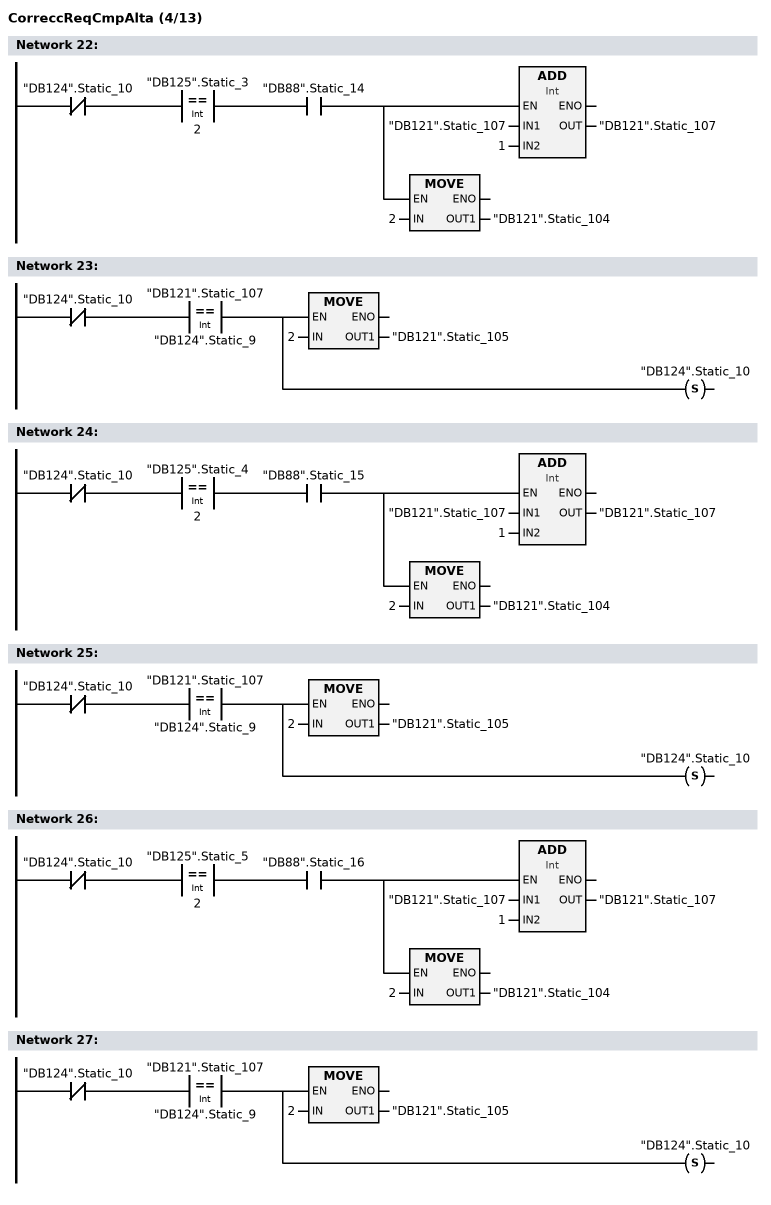
   IF NOT "DB124".Static_10 AND ("DB125".Static_3 = 2) AND "DB88".Static_14 THEN
       "DB121".Static_107 := "DB121".Static_107 + 1;
       "DB121".Static_104 := 2;
   END_IF;
END_REGION

REGION Network 23
   IF NOT "DB124".Static_10 AND ("DB121".Static_107 = "DB124".Static_9) THEN
       "DB121".Static_105 := 2;
       "DB124".Static_10 := TRUE;
   END_IF;
END_REGION

REGION Network 24
   IF NOT "DB124".Static_10 AND ("DB125".Static_4 = 2) AND "DB88".Static_15 THEN
       "DB121".Static_107 := "DB121".Static_107 + 1;
       "DB121".Static_104 := 2;
   END_IF;
END_REGION

REGION Network 25
   IF NOT "DB124".Static_10 AND ("DB121".Static_107 = "DB124".Static_9) THEN
       "DB121".Static_105 := 2;
       "DB124".Static_10 := TRUE;
   END_IF;
END_REGION

REGION Network 26
   IF NOT "DB124".Static_10 AND ("DB125".Static_5 = 2) AND "DB88".Static_16 THEN
       "DB121".Static_107 := "DB121".Static_107 + 1;
       "DB121".Static_104 := 2;
   END_IF;
END_REGION

REGION Network 27
   IF NOT "DB124".Static_10 AND ("DB121".Static_107 = "DB124".Static_9) THEN
       "DB121".Static_105 := 2;
       "DB124".Static_10 := TRUE;
   END_IF;
END_REGION

REGION Network 28
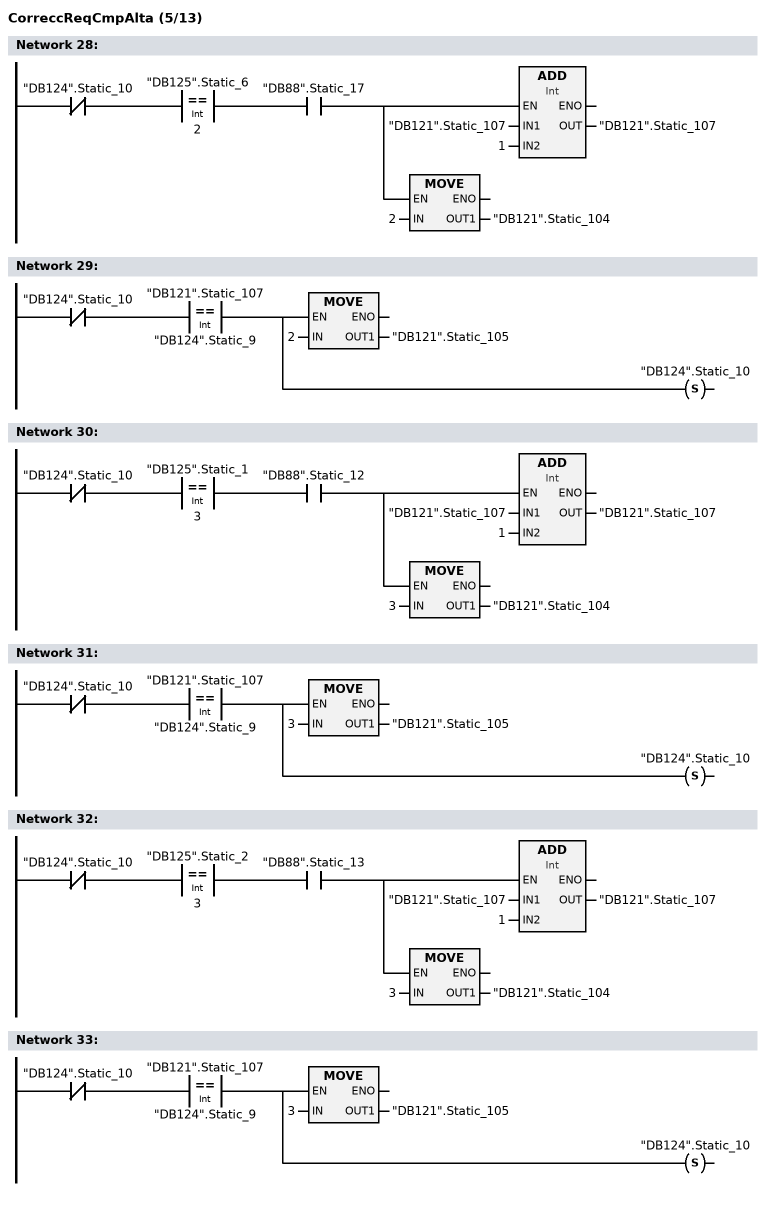
   IF NOT "DB124".Static_10 AND ("DB125".Static_6 = 2) AND "DB88".Static_17 THEN
       "DB121".Static_107 := "DB121".Static_107 + 1;
       "DB121".Static_104 := 2;
   END_IF;
END_REGION

REGION Network 29
   IF NOT "DB124".Static_10 AND ("DB121".Static_107 = "DB124".Static_9) THEN
       "DB121".Static_105 := 2;
       "DB124".Static_10 := TRUE;
   END_IF;
END_REGION

REGION Network 30
   IF NOT "DB124".Static_10 AND ("DB125".Static_1 = 3) AND "DB88".Static_12 THEN
       "DB121".Static_107 := "DB121".Static_107 + 1;
       "DB121".Static_104 := 3;
   END_IF;
END_REGION

REGION Network 31
   IF NOT "DB124".Static_10 AND ("DB121".Static_107 = "DB124".Static_9) THEN
       "DB121".Static_105 := 3;
       "DB124".Static_10 := TRUE;
   END_IF;
END_REGION

REGION Network 32
   IF NOT "DB124".Static_10 AND ("DB125".Static_2 = 3) AND "DB88".Static_13 THEN
       "DB121".Static_107 := "DB121".Static_107 + 1;
       "DB121".Static_104 := 3;
   END_IF;
END_REGION

REGION Network 33
   IF NOT "DB124".Static_10 AND ("DB121".Static_107 = "DB124".Static_9) THEN
       "DB121".Static_105 := 3;
       "DB124".Static_10 := TRUE;
   END_IF;
END_REGION

REGION Network 34
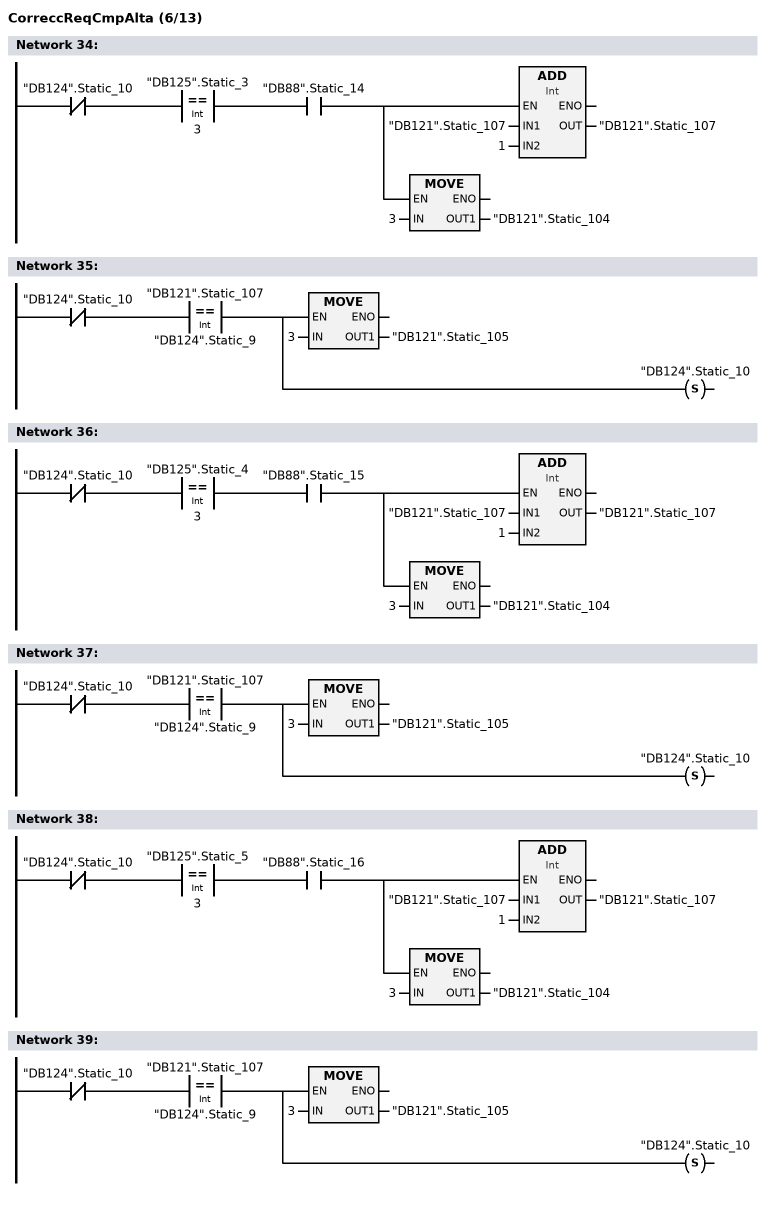
   IF NOT "DB124".Static_10 AND ("DB125".Static_3 = 3) AND "DB88".Static_14 THEN
       "DB121".Static_107 := "DB121".Static_107 + 1;
       "DB121".Static_104 := 3;
   END_IF;
END_REGION

REGION Network 35
   IF NOT "DB124".Static_10 AND ("DB121".Static_107 = "DB124".Static_9) THEN
       "DB121".Static_105 := 3;
       "DB124".Static_10 := TRUE;
   END_IF;
END_REGION

REGION Network 36
   IF NOT "DB124".Static_10 AND ("DB125".Static_4 = 3) AND "DB88".Static_15 THEN
       "DB121".Static_107 := "DB121".Static_107 + 1;
       "DB121".Static_104 := 3;
   END_IF;
END_REGION

REGION Network 37
   IF NOT "DB124".Static_10 AND ("DB121".Static_107 = "DB124".Static_9) THEN
       "DB121".Static_105 := 3;
       "DB124".Static_10 := TRUE;
   END_IF;
END_REGION

REGION Network 38
   IF NOT "DB124".Static_10 AND ("DB125".Static_5 = 3) AND "DB88".Static_16 THEN
       "DB121".Static_107 := "DB121".Static_107 + 1;
       "DB121".Static_104 := 3;
   END_IF;
END_REGION

REGION Network 39
   IF NOT "DB124".Static_10 AND ("DB121".Static_107 = "DB124".Static_9) THEN
       "DB121".Static_105 := 3;
       "DB124".Static_10 := TRUE;
   END_IF;
END_REGION

REGION Network 40
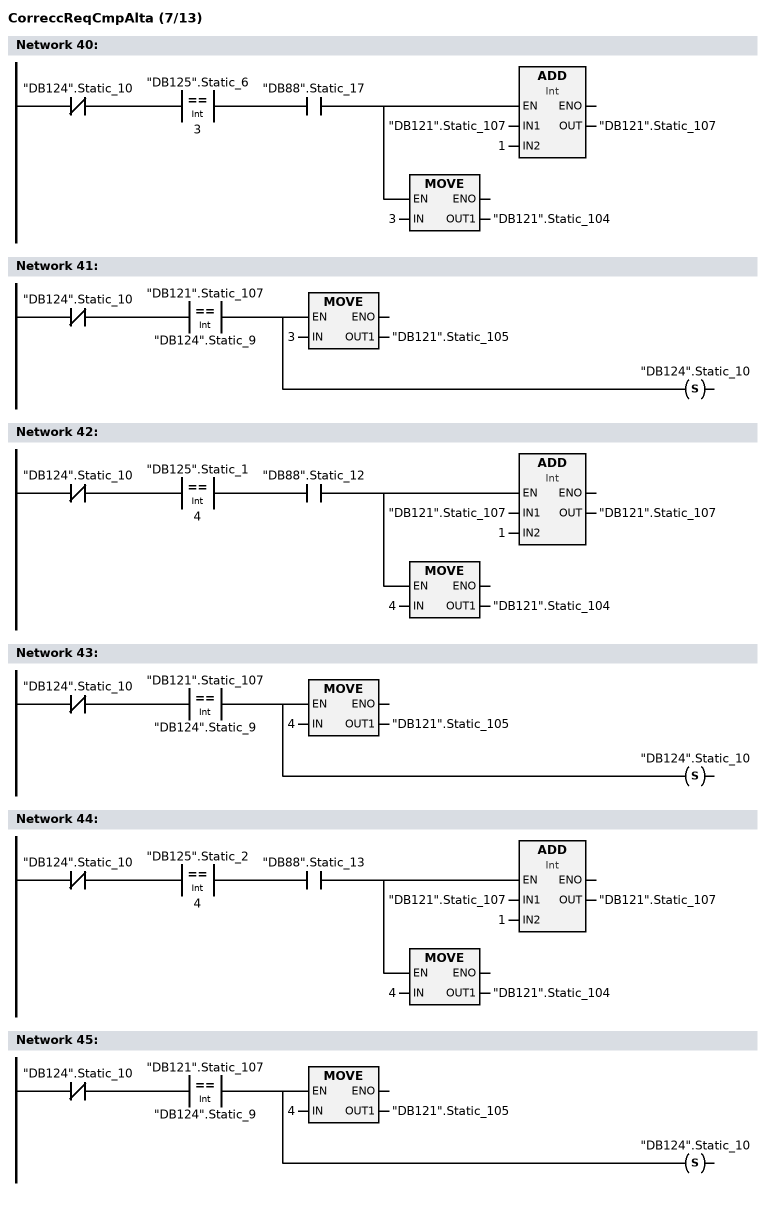
   IF NOT "DB124".Static_10 AND ("DB125".Static_6 = 3) AND "DB88".Static_17 THEN
       "DB121".Static_107 := "DB121".Static_107 + 1;
       "DB121".Static_104 := 3;
   END_IF;
END_REGION

REGION Network 41
   IF NOT "DB124".Static_10 AND ("DB121".Static_107 = "DB124".Static_9) THEN
       "DB121".Static_105 := 3;
       "DB124".Static_10 := TRUE;
   END_IF;
END_REGION

REGION Network 42
   IF NOT "DB124".Static_10 AND ("DB125".Static_1 = 4) AND "DB88".Static_12 THEN
       "DB121".Static_107 := "DB121".Static_107 + 1;
       "DB121".Static_104 := 4;
   END_IF;
END_REGION

REGION Network 43
   IF NOT "DB124".Static_10 AND ("DB121".Static_107 = "DB124".Static_9) THEN
       "DB121".Static_105 := 4;
       "DB124".Static_10 := TRUE;
   END_IF;
END_REGION

REGION Network 44
   IF NOT "DB124".Static_10 AND ("DB125".Static_2 = 4) AND "DB88".Static_13 THEN
       "DB121".Static_107 := "DB121".Static_107 + 1;
       "DB121".Static_104 := 4;
   END_IF;
END_REGION

REGION Network 45
   IF NOT "DB124".Static_10 AND ("DB121".Static_107 = "DB124".Static_9) THEN
       "DB121".Static_105 := 4;
       "DB124".Static_10 := TRUE;
   END_IF;
END_REGION

REGION Network 46
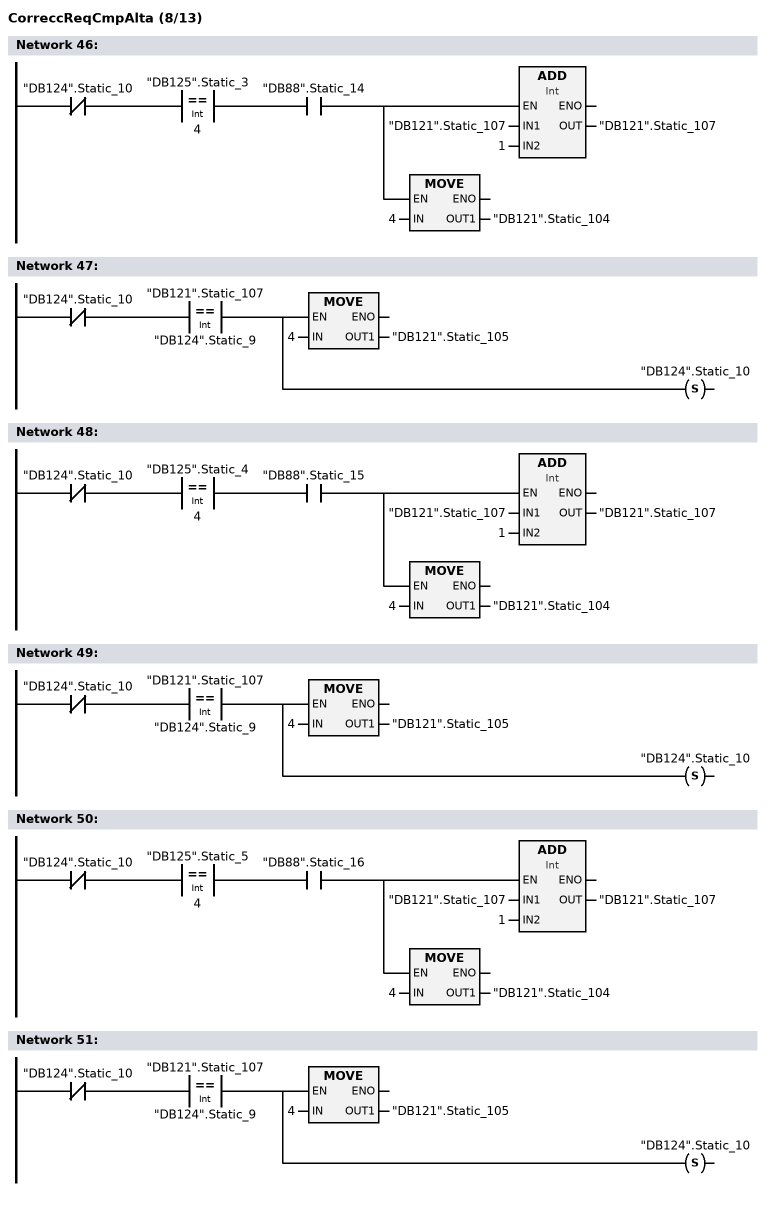
   IF NOT "DB124".Static_10 AND ("DB125".Static_3 = 4) AND "DB88".Static_14 THEN
       "DB121".Static_107 := "DB121".Static_107 + 1;
       "DB121".Static_104 := 4;
   END_IF;
END_REGION

REGION Network 47
   IF NOT "DB124".Static_10 AND ("DB121".Static_107 = "DB124".Static_9) THEN
       "DB121".Static_105 := 4;
       "DB124".Static_10 := TRUE;
   END_IF;
END_REGION

REGION Network 48
   IF NOT "DB124".Static_10 AND ("DB125".Static_4 = 4) AND "DB88".Static_15 THEN
       "DB121".Static_107 := "DB121".Static_107 + 1;
       "DB121".Static_104 := 4;
   END_IF;
END_REGION

REGION Network 49
   IF NOT "DB124".Static_10 AND ("DB121".Static_107 = "DB124".Static_9) THEN
       "DB121".Static_105 := 4;
       "DB124".Static_10 := TRUE;
   END_IF;
END_REGION

REGION Network 50
   IF NOT "DB124".Static_10 AND ("DB125".Static_5 = 4) AND "DB88".Static_16 THEN
       "DB121".Static_107 := "DB121".Static_107 + 1;
       "DB121".Static_104 := 4;
   END_IF;
END_REGION

REGION Network 51
   IF NOT "DB124".Static_10 AND ("DB121".Static_107 = "DB124".Static_9) THEN
       "DB121".Static_105 := 4;
       "DB124".Static_10 := TRUE;
   END_IF;
END_REGION

REGION Network 52
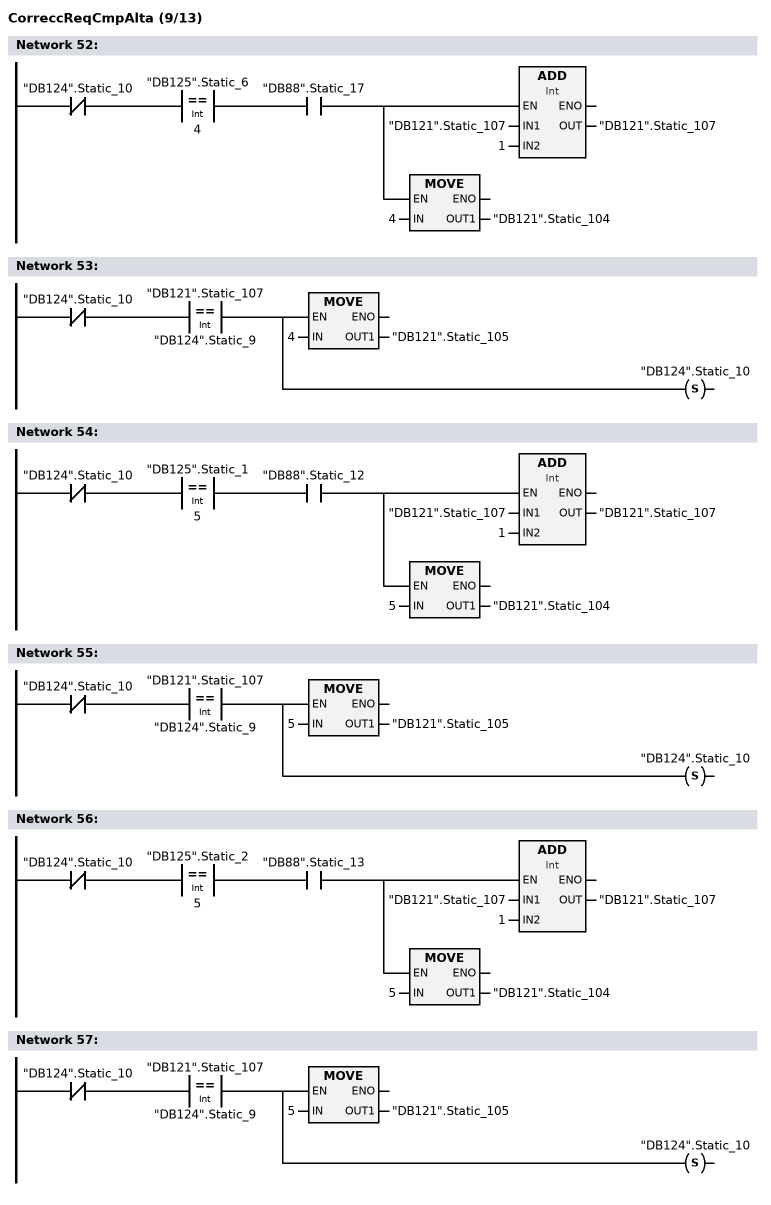
   IF NOT "DB124".Static_10 AND ("DB125".Static_6 = 4) AND "DB88".Static_17 THEN
       "DB121".Static_107 := "DB121".Static_107 + 1;
       "DB121".Static_104 := 4;
   END_IF;
END_REGION

REGION Network 53
   IF NOT "DB124".Static_10 AND ("DB121".Static_107 = "DB124".Static_9) THEN
       "DB121".Static_105 := 4;
       "DB124".Static_10 := TRUE;
   END_IF;
END_REGION

REGION Network 54
   IF NOT "DB124".Static_10 AND ("DB125".Static_1 = 5) AND "DB88".Static_12 THEN
       "DB121".Static_107 := "DB121".Static_107 + 1;
       "DB121".Static_104 := 5;
   END_IF;
END_REGION

REGION Network 55
   IF NOT "DB124".Static_10 AND ("DB121".Static_107 = "DB124".Static_9) THEN
       "DB121".Static_105 := 5;
       "DB124".Static_10 := TRUE;
   END_IF;
END_REGION

REGION Network 56
   IF NOT "DB124".Static_10 AND ("DB125".Static_2 = 5) AND "DB88".Static_13 THEN
       "DB121".Static_107 := "DB121".Static_107 + 1;
       "DB121".Static_104 := 5;
   END_IF;
END_REGION

REGION Network 57
   IF NOT "DB124".Static_10 AND ("DB121".Static_107 = "DB124".Static_9) THEN
       "DB121".Static_105 := 5;
       "DB124".Static_10 := TRUE;
   END_IF;
END_REGION

REGION Network 58
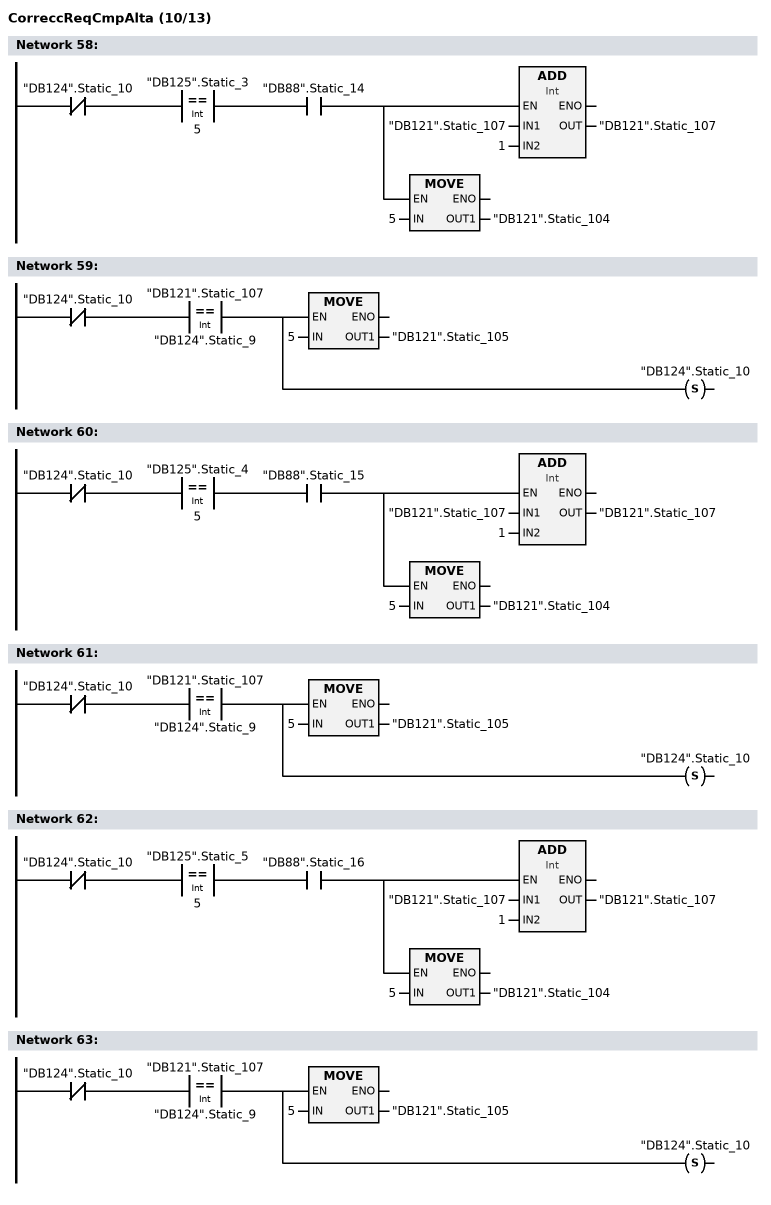
   IF NOT "DB124".Static_10 AND ("DB125".Static_3 = 5) AND "DB88".Static_14 THEN
       "DB121".Static_107 := "DB121".Static_107 + 1;
       "DB121".Static_104 := 5;
   END_IF;
END_REGION

REGION Network 59
   IF NOT "DB124".Static_10 AND ("DB121".Static_107 = "DB124".Static_9) THEN
       "DB121".Static_105 := 5;
       "DB124".Static_10 := TRUE;
   END_IF;
END_REGION

REGION Network 60
   IF NOT "DB124".Static_10 AND ("DB125".Static_4 = 5) AND "DB88".Static_15 THEN
       "DB121".Static_107 := "DB121".Static_107 + 1;
       "DB121".Static_104 := 5;
   END_IF;
END_REGION

REGION Network 61
   IF NOT "DB124".Static_10 AND ("DB121".Static_107 = "DB124".Static_9) THEN
       "DB121".Static_105 := 5;
       "DB124".Static_10 := TRUE;
   END_IF;
END_REGION

REGION Network 62
   IF NOT "DB124".Static_10 AND ("DB125".Static_5 = 5) AND "DB88".Static_16 THEN
       "DB121".Static_107 := "DB121".Static_107 + 1;
       "DB121".Static_104 := 5;
   END_IF;
END_REGION

REGION Network 63
   IF NOT "DB124".Static_10 AND ("DB121".Static_107 = "DB124".Static_9) THEN
       "DB121".Static_105 := 5;
       "DB124".Static_10 := TRUE;
   END_IF;
END_REGION

REGION Network 64
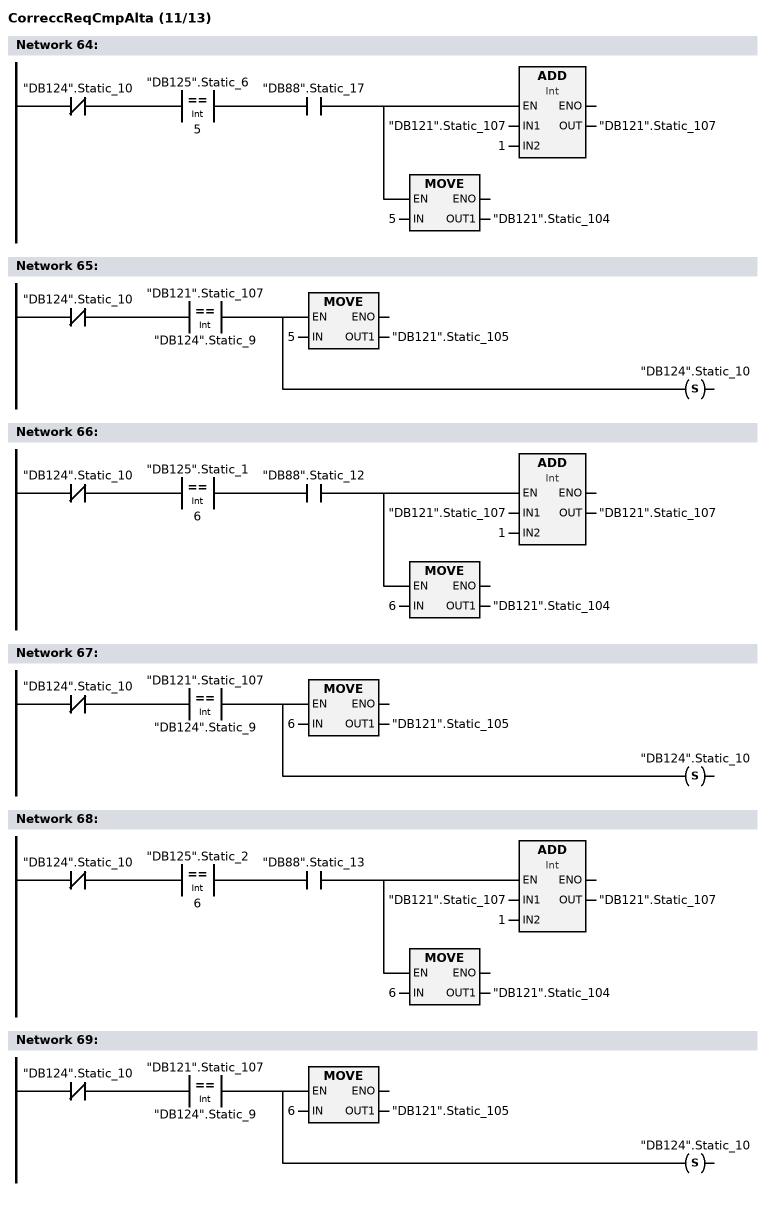
   IF NOT "DB124".Static_10 AND ("DB125".Static_6 = 5) AND "DB88".Static_17 THEN
       "DB121".Static_107 := "DB121".Static_107 + 1;
       "DB121".Static_104 := 5;
   END_IF;
END_REGION

REGION Network 65
   IF NOT "DB124".Static_10 AND ("DB121".Static_107 = "DB124".Static_9) THEN
       "DB121".Static_105 := 5;
       "DB124".Static_10 := TRUE;
   END_IF;
END_REGION

REGION Network 66
   IF NOT "DB124".Static_10 AND ("DB125".Static_1 = 6) AND "DB88".Static_12 THEN
       "DB121".Static_107 := "DB121".Static_107 + 1;
       "DB121".Static_104 := 6;
   END_IF;
END_REGION

REGION Network 67
   IF NOT "DB124".Static_10 AND ("DB121".Static_107 = "DB124".Static_9) THEN
       "DB121".Static_105 := 6;
       "DB124".Static_10 := TRUE;
   END_IF;
END_REGION

REGION Network 68
   IF NOT "DB124".Static_10 AND ("DB125".Static_2 = 6) AND "DB88".Static_13 THEN
       "DB121".Static_107 := "DB121".Static_107 + 1;
       "DB121".Static_104 := 6;
   END_IF;
END_REGION

REGION Network 69
   IF NOT "DB124".Static_10 AND ("DB121".Static_107 = "DB124".Static_9) THEN
       "DB121".Static_105 := 6;
       "DB124".Static_10 := TRUE;
   END_IF;
END_REGION

REGION Network 70
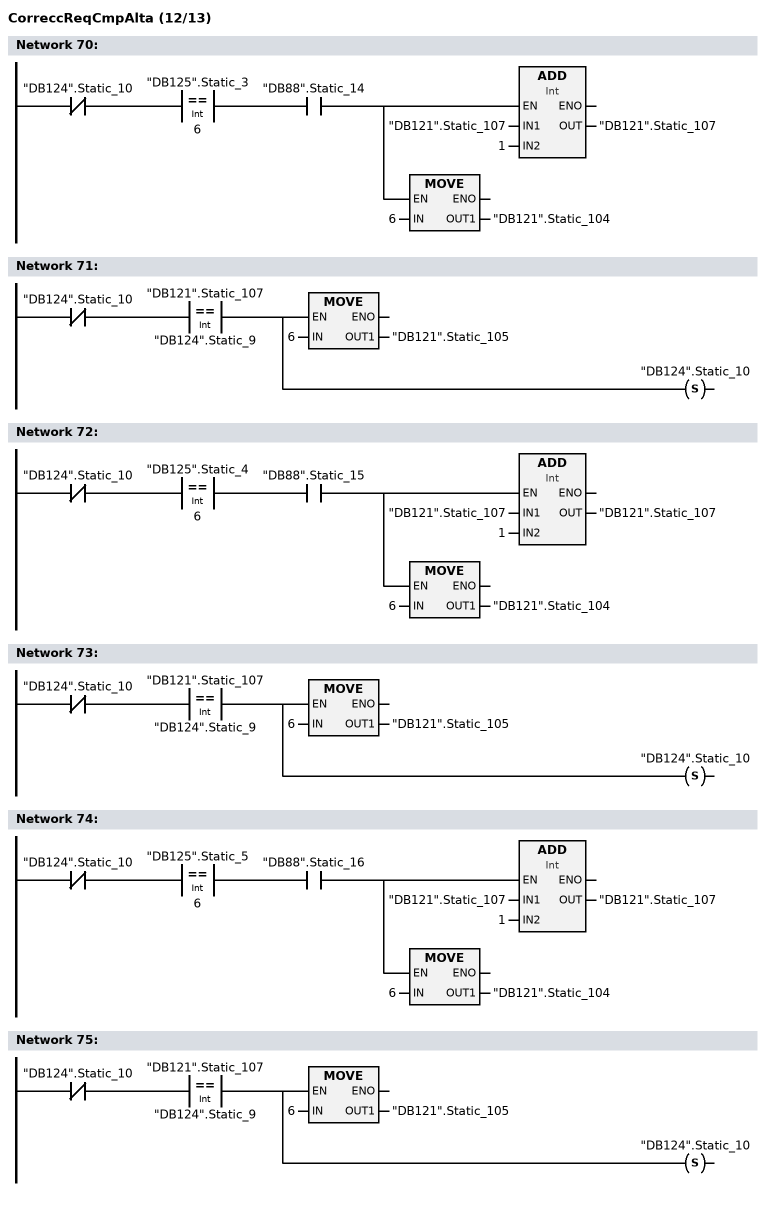
   IF NOT "DB124".Static_10 AND ("DB125".Static_3 = 6) AND "DB88".Static_14 THEN
       "DB121".Static_107 := "DB121".Static_107 + 1;
       "DB121".Static_104 := 6;
   END_IF;
END_REGION

REGION Network 71
   IF NOT "DB124".Static_10 AND ("DB121".Static_107 = "DB124".Static_9) THEN
       "DB121".Static_105 := 6;
       "DB124".Static_10 := TRUE;
   END_IF;
END_REGION

REGION Network 72
   IF NOT "DB124".Static_10 AND ("DB125".Static_4 = 6) AND "DB88".Static_15 THEN
       "DB121".Static_107 := "DB121".Static_107 + 1;
       "DB121".Static_104 := 6;
   END_IF;
END_REGION

REGION Network 73
   IF NOT "DB124".Static_10 AND ("DB121".Static_107 = "DB124".Static_9) THEN
       "DB121".Static_105 := 6;
       "DB124".Static_10 := TRUE;
   END_IF;
END_REGION

REGION Network 74
   IF NOT "DB124".Static_10 AND ("DB125".Static_5 = 6) AND "DB88".Static_16 THEN
       "DB121".Static_107 := "DB121".Static_107 + 1;
       "DB121".Static_104 := 6;
   END_IF;
END_REGION

REGION Network 75
   IF NOT "DB124".Static_10 AND ("DB121".Static_107 = "DB124".Static_9) THEN
       "DB121".Static_105 := 6;
       "DB124".Static_10 := TRUE;
   END_IF;
END_REGION

REGION Network 76
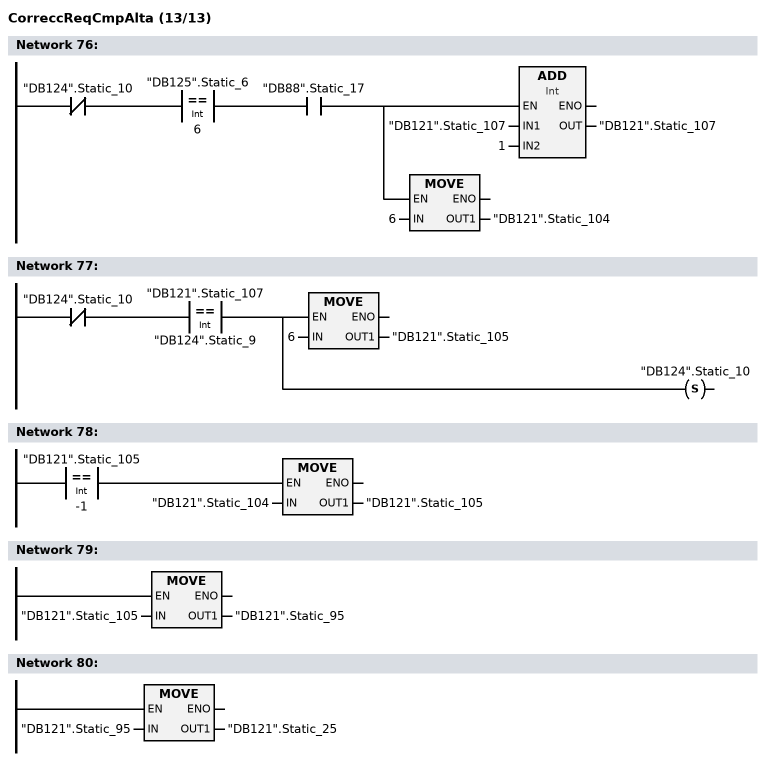
   IF NOT "DB124".Static_10 AND ("DB125".Static_6 = 6) AND "DB88".Static_17 THEN
       "DB121".Static_107 := "DB121".Static_107 + 1;
       "DB121".Static_104 := 6;
   END_IF;
END_REGION

REGION Network 77
   IF NOT "DB124".Static_10 AND ("DB121".Static_107 = "DB124".Static_9) THEN
       "DB121".Static_105 := 6;
       "DB124".Static_10 := TRUE;
   END_IF;
END_REGION

REGION Network 78
   RUNG wire#powerrail
      { S7_Templates := "SrcType := Int" } EQ_Contact(in1 := "DB121".Static_105, in2 := -1)
      { S7_GenerateENO := "TRUE" } Move(in := "DB121".Static_104, out1 => "DB121".Static_105)
   END_RUNG
   // the same network as SCL:
   IF "DB121".Static_105 = (-1) THEN "DB121".Static_105 := "DB121".Static_104; END_IF;
END_REGION

REGION Network 79
   RUNG wire#powerrail
      { S7_GenerateENO := "TRUE" } Move(in := "DB121".Static_105, out1 => "DB121".Static_95)
   END_RUNG
   // the same network as SCL:
   "DB121".Static_95 := "DB121".Static_105;
END_REGION

REGION Network 80
   RUNG wire#powerrail
      { S7_GenerateENO := "TRUE" } Move(in := "DB121".Static_95, out1 => "DB121".Static_25)
   END_RUNG
   // the same network as SCL:
   "DB121".Static_25 := "DB121".Static_95;
END_REGION
END_FUNCTION

FUNCTION "CalcEst6" : Void   // FC50, LAD
{ S7_Optimized_Access := 'FALSE' }
VERSION : 0.1
   VAR_TEMP   // added for the SCL form of the ladder/FBD networks
      _w1 : Bool;
   END_VAR
BEGIN

REGION Network 1
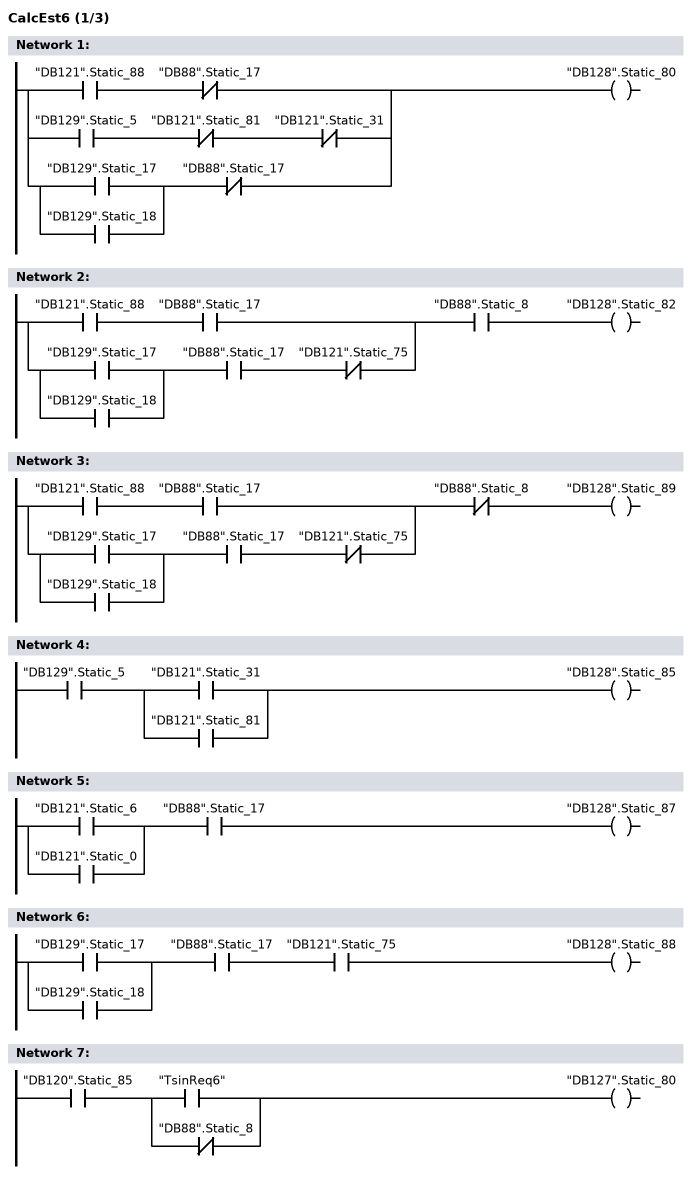
   RUNG wire#powerrail
      Contact( "DB121".Static_88 )
      I_Contact( "DB88".Static_17 )
      wire#w1
      Coil( "DB128".Static_80 )
   END_RUNG
   RUNG wire#powerrail
      Contact( "DB129".Static_5 )
      I_Contact( "DB121".Static_81 )
      I_Contact( "DB121".Static_31 )
   END_RUNG wire#w1
   RUNG wire#powerrail
      Contact( "DB129".Static_17 )
      wire#w2
      I_Contact( "DB88".Static_17 )
   END_RUNG wire#w1
   RUNG wire#powerrail
      Contact( "DB129".Static_18 )
   END_RUNG wire#w2
   // the same network as SCL:
   "DB128".Static_80 := ("DB121".Static_88 AND NOT "DB88".Static_17) OR ("DB129".Static_5 AND NOT "DB121".Static_81 AND NOT "DB121".Static_31) OR (("DB129".Static_17 OR "DB129".Static_18) AND NOT "DB88".Static_17);
END_REGION

REGION Network 2
   RUNG wire#powerrail
      Contact( "DB121".Static_88 )
      Contact( "DB88".Static_17 )
      wire#w1
      Contact( "DB88".Static_8 )
      Coil( "DB128".Static_82 )
   END_RUNG
   RUNG wire#powerrail
      Contact( "DB129".Static_17 )
      wire#w2
      Contact( "DB88".Static_17 )
      I_Contact( "DB121".Static_75 )
   END_RUNG wire#w1
   RUNG wire#powerrail
      Contact( "DB129".Static_18 )
   END_RUNG wire#w2
   // the same network as SCL:
   "DB128".Static_82 := (("DB121".Static_88 AND "DB88".Static_17) OR (("DB129".Static_17 OR "DB129".Static_18) AND "DB88".Static_17 AND NOT "DB121".Static_75)) AND "DB88".Static_8;
END_REGION

REGION Network 3
   RUNG wire#powerrail
      Contact( "DB121".Static_88 )
      Contact( "DB88".Static_17 )
      wire#w1
      I_Contact( "DB88".Static_8 )
      Coil( "DB128".Static_89 )
   END_RUNG
   RUNG wire#powerrail
      Contact( "DB129".Static_17 )
      wire#w2
      Contact( "DB88".Static_17 )
      I_Contact( "DB121".Static_75 )
   END_RUNG wire#w1
   RUNG wire#powerrail
      Contact( "DB129".Static_18 )
   END_RUNG wire#w2
   // the same network as SCL:
   "DB128".Static_89 := (("DB121".Static_88 AND "DB88".Static_17) OR (("DB129".Static_17 OR "DB129".Static_18) AND "DB88".Static_17 AND NOT "DB121".Static_75)) AND NOT "DB88".Static_8;
END_REGION

REGION Network 4
   "DB128".Static_85 := "DB129".Static_5 AND ("DB121".Static_31 OR "DB121".Static_81);
END_REGION

REGION Network 5
   RUNG wire#powerrail
      Contact( "DB121".Static_6 )
      wire#w1
      Contact( "DB88".Static_17 )
      Coil( "DB128".Static_87 )
   END_RUNG
   RUNG wire#powerrail
      Contact( "DB121".Static_0 )
   END_RUNG wire#w1
   // the same network as SCL:
   "DB128".Static_87 := ("DB121".Static_6 OR "DB121".Static_0) AND "DB88".Static_17;
END_REGION

REGION Network 6
   RUNG wire#powerrail
      Contact( "DB129".Static_17 )
      wire#w1
      Contact( "DB88".Static_17 )
      Contact( "DB121".Static_75 )
      Coil( "DB128".Static_88 )
   END_RUNG
   RUNG wire#powerrail
      Contact( "DB129".Static_18 )
   END_RUNG wire#w1
   // the same network as SCL:
   "DB128".Static_88 := ("DB129".Static_17 OR "DB129".Static_18) AND "DB88".Static_17 AND "DB121".Static_75;
END_REGION

REGION Network 7
   "DB127".Static_80 := "DB120".Static_85 AND ("TsinReq6" OR NOT "DB88".Static_8);
END_REGION

REGION Network 8
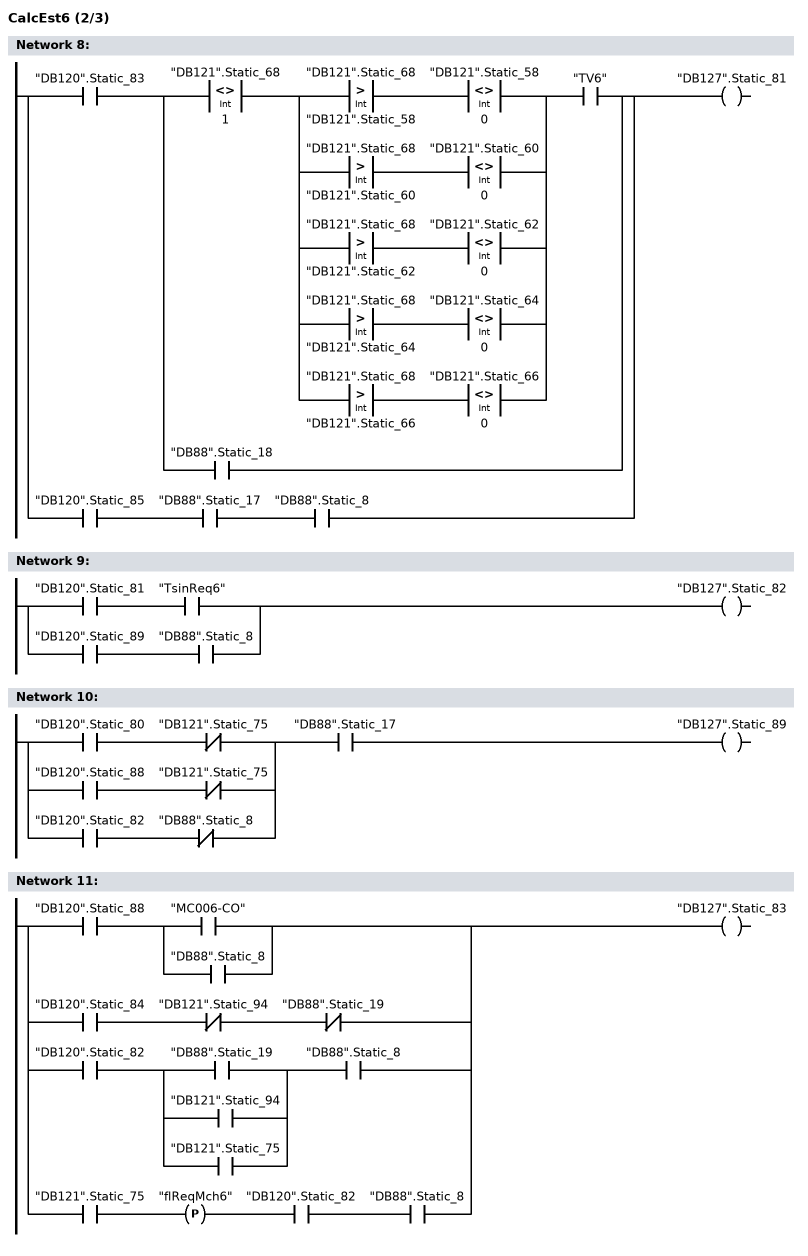
   "DB127".Static_81 := ("DB120".Static_83 AND ((("DB121".Static_68 <> 1) AND ((("DB121".Static_68 > "DB121".Static_58) AND ("DB121".Static_58 <> 0)) OR (("DB121".Static_68 > "DB121".Static_60) AND ("DB121".Static_60 <> 0)) OR (("DB121".Static_68 > "DB121".Static_62) AND ("DB121".Static_62 <> 0)) OR (("DB121".Static_68 > "DB121".Static_64) AND ("DB121".Static_64 <> 0)) OR (("DB121".Static_68 > "DB121".Static_66) AND ("DB121".Static_66 <> 0))) AND "TV6") OR "DB88".Static_18)) OR ("DB120".Static_85 AND "DB88".Static_17 AND "DB88".Static_8);
END_REGION
